// TIA Portal project "Sistema_de_silos" (V16) (continued)
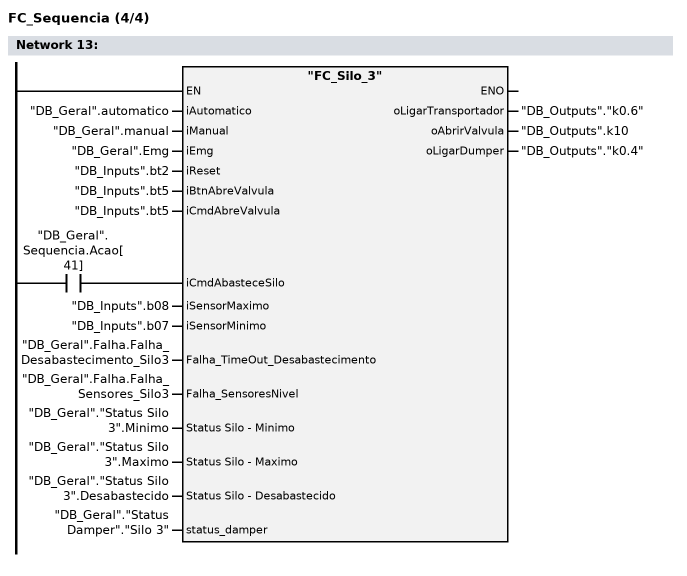
   RUNG wire#powerrail
      "FC_Silo_3"(iCmdAbasteceSilo := wire#w1, iAutomatico := "DB_Geral".automatico, iManual := "DB_Geral".manual, iEmg := "DB_Geral".Emg, iReset := "DB_Inputs".bt2, iBtnAbreValvula := "DB_Inputs".bt5, iCmdAbreValvula := "DB_Inputs".bt5, iSensorMaximo := "DB_Inputs".b08, iSensorMinimo := "DB_Inputs".b07, Falha_TimeOut_Desabastecimento := "DB_Geral".Falha.Falha_Desabastecimento_Silo3, Falha_SensoresNivel := "DB_Geral".Falha.Falha_Sensores_Silo3, "Status Silo - Minimo" := "DB_Geral"."Status Silo 3".Minimo, "Status Silo - Maximo" := "DB_Geral"."Status Silo 3".Maximo, "Status Silo - Desabastecido" := "DB_Geral"."Status Silo 3".Desabastecido, status_damper := "DB_Geral"."Status Damper"."Silo 3", oLigarTransportador => "DB_Outputs"."k0.6", oAbrirValvula => "DB_Outputs".k10, oLigarDumper => "DB_Outputs"."k0.4")
   END_RUNG
   RUNG wire#powerrail
      Contact( "DB_Geral".Sequencia.Acao[41] )
   END_RUNG wire#w1
   // the same network as SCL:
   "FC_Silo_3"(iAutomatico := "DB_Geral".automatico,
               iManual := "DB_Geral".manual,
               iEmg := "DB_Geral".Emg,
               iReset := "DB_Inputs".bt2,
               iBtnAbreValvula := "DB_Inputs".bt5,
               iCmdAbreValvula := "DB_Inputs".bt5,
               iCmdAbasteceSilo := "DB_Geral".Sequencia.Acao[41],
               iSensorMaximo := "DB_Inputs".b08,
               iSensorMinimo := "DB_Inputs".b07,
               Falha_TimeOut_Desabastecimento := "DB_Geral".Falha.Falha_Desabastecimento_Silo3,
               Falha_SensoresNivel := "DB_Geral".Falha.Falha_Sensores_Silo3,
               "Status Silo - Minimo" := "DB_Geral"."Status Silo 3".Minimo,
               "Status Silo - Maximo" := "DB_Geral"."Status Silo 3".Maximo,
               "Status Silo - Desabastecido" := "DB_Geral"."Status Silo 3".Desabastecido,
               status_damper := "DB_Geral"."Status Damper"."Silo 3",
               oLigarTransportador => "DB_Outputs"."k0.6",
               oAbrirValvula => "DB_Outputs".k10,
               oLigarDumper => "DB_Outputs"."k0.4");
END_REGION
END_FUNCTION

FUNCTION "FC_Silo_2" : Void   // FC5, LAD
{ S7_Optimized_Access := 'TRUE' }
VERSION : 0.1
   VAR_INPUT
      iAutomatico : Bool;
      iManual : Bool;
      iEmg : Bool;
      iReset : Bool;
      iBtnAbreValvula : Bool;
      iCmdAbreValvula : Bool;
      iCmdAbasteceSilo : Bool;
      iSensorMaximo : Bool;
      iSensorMinimo : Bool;
   END_VAR
   VAR_OUTPUT
      oLigarTransportador : Bool;
      oAbrirValvula : Bool;
      oLigarDumper : Bool;
   END_VAR
   VAR_IN_OUT
      Falha_TimeOut_Desabastecimento : Bool;
      Falha_SensoresNivel : Bool;
      "Status Silo - Minimo" : Bool;
      "Status Silo - Maximo" : Bool;
      "Status Silo - Desabastecido" : Bool;
      status_damper : Bool;
   END_VAR
   VAR CONSTANT
      Velocidade_fluxo : Int := 12;
   END_VAR
BEGIN

REGION Network 1
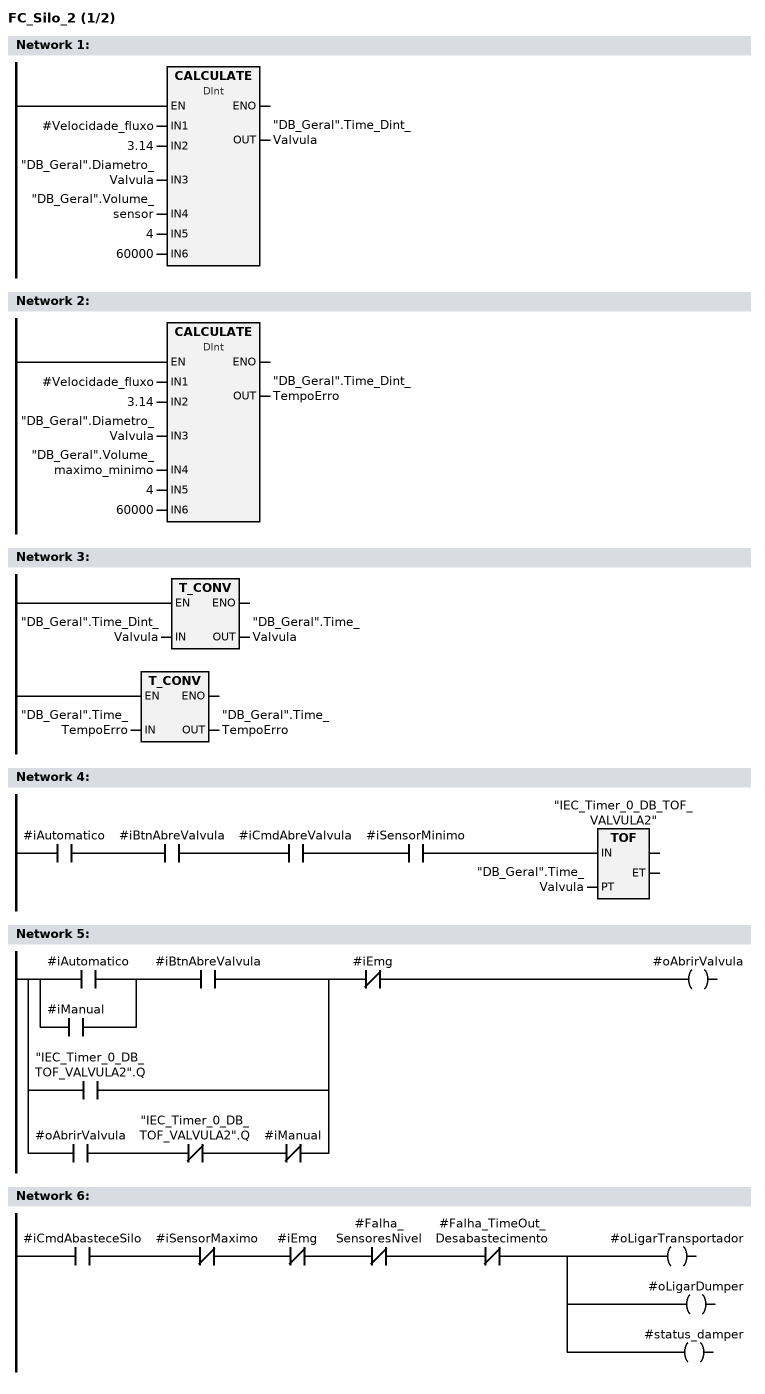
   RUNG wire#powerrail
      { S7_Templates := "SrcType := DInt"; S7_Expression := "(IN4 / (IN1* ((IN2*IN3*IN3) / IN5))) * IN6" } Calculate(in1 := #Velocidade_fluxo, in2 := 3.14, in3 := "DB_Geral".Diametro_Valvula, in4 := "DB_Geral".Volume_sensor, in5 := 4, in6 := 60000, out => "DB_Geral".Time_Dint_Valvula)
   END_RUNG
   // the same network as SCL:
   "DB_Geral".Time_Dint_Valvula := ("DB_Geral".Volume_sensor / (#Velocidade_fluxo* ((3.14*"DB_Geral".Diametro_Valvula*"DB_Geral".Diametro_Valvula) / 4))) * 60000;
END_REGION

REGION Network 2
   RUNG wire#powerrail
      { S7_Templates := "SrcType := DInt"; S7_Expression := "(IN4 / (IN1* ((IN2*IN3*IN3) / IN5))) * IN6" } Calculate(in1 := #Velocidade_fluxo, in2 := 3.14, in3 := "DB_Geral".Diametro_Valvula, in4 := "DB_Geral".Volume_maximo_minimo, in5 := 4, in6 := 60000, out => "DB_Geral".Time_Dint_TempoErro)
   END_RUNG
   // the same network as SCL:
   "DB_Geral".Time_Dint_TempoErro := ("DB_Geral".Volume_maximo_minimo / (#Velocidade_fluxo* ((3.14*"DB_Geral".Diametro_Valvula*"DB_Geral".Diametro_Valvula) / 4))) * 60000;
END_REGION

REGION Network 3
   "DB_Geral".Time_Valvula := T_CONV(IN := "DB_Geral".Time_Dint_Valvula);
   "DB_Geral".Time_TempoErro := T_CONV(IN := "DB_Geral".Time_TempoErro);
END_REGION

REGION Network 4
   "IEC_Timer_0_DB_TOF_VALVULA2".TOF(IN := #iAutomatico AND #iBtnAbreValvula AND #iCmdAbreValvula AND #iSensorMinimo,
                           PT := "DB_Geral".Time_Valvula);
END_REGION

REGION Network 5
   RUNG wire#powerrail
      Contact( #iAutomatico )
      wire#w1
      Contact( #iBtnAbreValvula )
      wire#w2
      I_Contact( #iEmg )
      Coil( #oAbrirValvula )
   END_RUNG
   RUNG wire#powerrail
      Contact( #iManual )
   END_RUNG wire#w1
   RUNG wire#powerrail
      Contact( "IEC_Timer_0_DB_TOF_VALVULA2".Q )
   END_RUNG wire#w2
   RUNG wire#powerrail
      Contact( #oAbrirValvula )
      I_Contact( "IEC_Timer_0_DB_TOF_VALVULA2".Q )
      I_Contact( #iManual )
   END_RUNG wire#w2
   // the same network as SCL:
   #oAbrirValvula := (((#iAutomatico OR #iManual) AND #iBtnAbreValvula) OR "IEC_Timer_0_DB_TOF_VALVULA2".Q OR (#oAbrirValvula AND NOT "IEC_Timer_0_DB_TOF_VALVULA2".Q AND NOT #iManual)) AND NOT #iEmg;
END_REGION

REGION Network 6
   RUNG wire#powerrail
      Contact( #iCmdAbasteceSilo )
      I_Contact( #iSensorMaximo )
      I_Contact( #iEmg )
      I_Contact( #Falha_SensoresNivel )
      I_Contact( #Falha_TimeOut_Desabastecimento )
      wire#w1
      Coil( #oLigarTransportador )
   END_RUNG
   RUNG wire#w1
      Coil( #oLigarDumper )
   END_RUNG
   RUNG wire#w1
      Coil( #status_damper )
   END_RUNG
   // the same network as SCL:
   #oLigarTransportador := #iCmdAbasteceSilo AND NOT #iSensorMaximo AND NOT #iEmg AND NOT #Falha_SensoresNivel AND NOT #Falha_TimeOut_Desabastecimento;
   #oLigarDumper := #oLigarTransportador;
   #status_damper := #oLigarTransportador;
END_REGION

REGION Network 7: Silo Principal - Reserva do produto
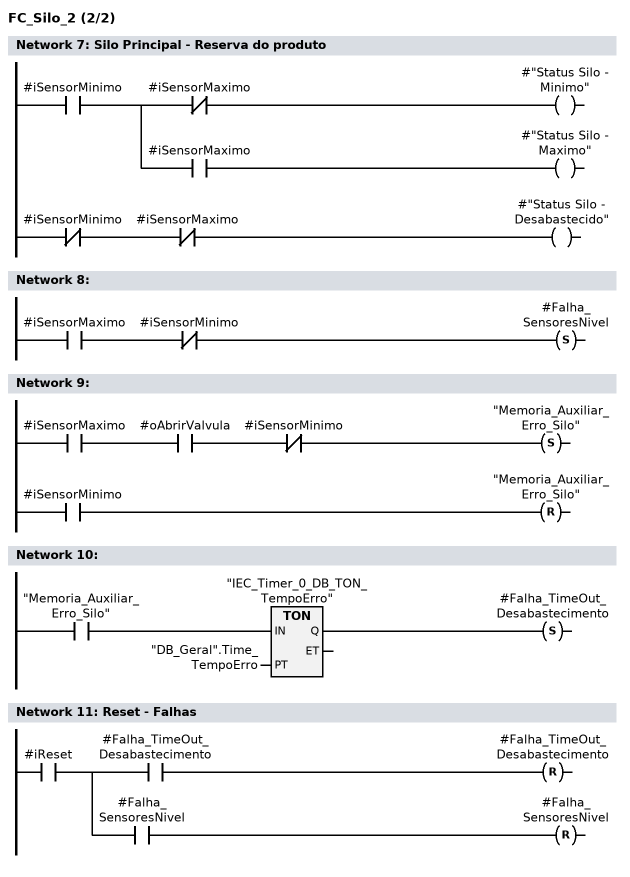
   RUNG wire#powerrail
      Contact( #iSensorMinimo )
      wire#w1
      I_Contact( #iSensorMaximo )
      Coil( #"Status Silo - Minimo" )
   END_RUNG
   RUNG wire#w1
      Contact( #iSensorMaximo )
      Coil( #"Status Silo - Maximo" )
   END_RUNG
   RUNG wire#powerrail
      I_Contact( #iSensorMinimo )
      I_Contact( #iSensorMaximo )
      Coil( #"Status Silo - Desabastecido" )
   END_RUNG
   // the same network as SCL:
   #"Status Silo - Minimo" := #iSensorMinimo AND NOT #iSensorMaximo;
   #"Status Silo - Maximo" := #iSensorMinimo AND #iSensorMaximo;
   #"Status Silo - Desabastecido" := NOT #iSensorMinimo AND NOT #iSensorMaximo;
END_REGION

REGION Network 8
   RUNG wire#powerrail
      Contact( #iSensorMaximo )
      I_Contact( #iSensorMinimo )
      S_Coil( #Falha_SensoresNivel )
   END_RUNG
   // the same network as SCL:
   IF #iSensorMaximo AND NOT #iSensorMinimo THEN #Falha_SensoresNivel := TRUE; END_IF;
END_REGION

REGION Network 9
   RUNG wire#powerrail
      Contact( #iSensorMaximo )
      Contact( #oAbrirValvula )
      I_Contact( #iSensorMinimo )
      S_Coil( "Memoria_Auxiliar_Erro_Silo" )
   END_RUNG
   RUNG wire#powerrail
      Contact( #iSensorMinimo )
      R_Coil( "Memoria_Auxiliar_Erro_Silo" )
   END_RUNG
   // the same network as SCL:
   IF #iSensorMaximo AND #oAbrirValvula AND NOT #iSensorMinimo THEN
       "Memoria_Auxiliar_Erro_Silo" := TRUE;
   END_IF;
   IF #iSensorMinimo THEN "Memoria_Auxiliar_Erro_Silo" := FALSE; END_IF;
END_REGION

REGION Network 10
   "IEC_Timer_0_DB_TON_TempoErro".TON(IN := "Memoria_Auxiliar_Erro_Silo", PT := "DB_Geral".Time_TempoErro);
   IF "IEC_Timer_0_DB_TON_TempoErro".Q THEN #Falha_TimeOut_Desabastecimento := TRUE; END_IF;
END_REGION

REGION Network 11: Reset - Falhas
   RUNG wire#powerrail
      Contact( #iReset )
      wire#w1
      Contact( #Falha_TimeOut_Desabastecimento )
      R_Coil( #Falha_TimeOut_Desabastecimento )
   END_RUNG
   RUNG wire#w1
      Contact( #Falha_SensoresNivel )
      R_Coil( #Falha_SensoresNivel )
   END_RUNG
   // the same network as SCL:
   IF #iReset AND #Falha_TimeOut_Desabastecimento THEN #Falha_TimeOut_Desabastecimento := FALSE; END_IF;
   IF #iReset AND #Falha_SensoresNivel THEN #Falha_SensoresNivel := FALSE; END_IF;
END_REGION
END_FUNCTION

FUNCTION "FC_Silo_Principal" : Void   // FC6, LAD
{ S7_Optimized_Access := 'TRUE' }
VERSION : 0.1
   VAR_INPUT
      iAutomatico : Bool;
      iManual : Bool;
      iEmg : Bool;
      iReset : Bool;
      iBtnAbasteceSilo : Bool;
      iCmdAbasteceSilo : Bool;
      iSensorMaximo : Bool;
      iSensorMinimo : Bool;
   END_VAR
   VAR_OUTPUT
      oAbasteceSilo : Bool;
   END_VAR
   VAR_IN_OUT
      Falha_SensoresNivel : Bool;
      "Status Silo - Minimo" : Bool;
      "Status Silo - Maximo" : Bool;
      "Status Silo - Desabastecido" : Bool;
   END_VAR
BEGIN

REGION Network 1
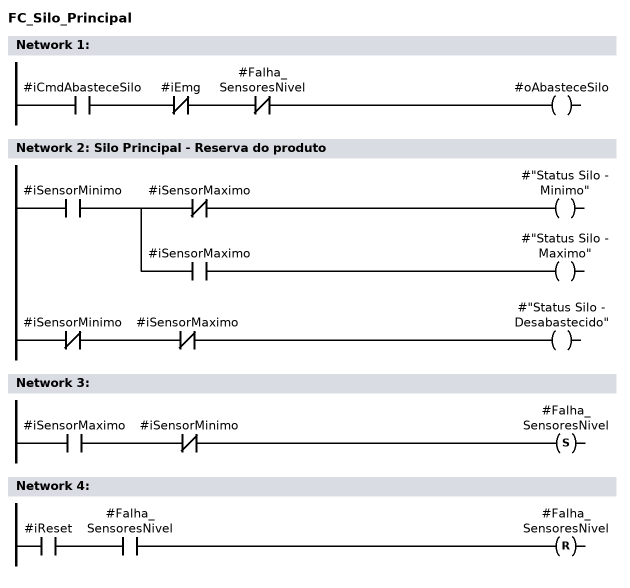
   RUNG wire#powerrail
      Contact( #iCmdAbasteceSilo )
      I_Contact( #iEmg )
      I_Contact( #Falha_SensoresNivel )
      Coil( #oAbasteceSilo )
   END_RUNG
   // the same network as SCL:
   #oAbasteceSilo := #iCmdAbasteceSilo AND NOT #iEmg AND NOT #Falha_SensoresNivel;
END_REGION

REGION Network 2: Silo Principal - Reserva do produto
   RUNG wire#powerrail
      Contact( #iSensorMinimo )
      wire#w1
      I_Contact( #iSensorMaximo )
      Coil( #"Status Silo - Minimo" )
   END_RUNG
   RUNG wire#w1
      Contact( #iSensorMaximo )
      Coil( #"Status Silo - Maximo" )
   END_RUNG
   RUNG wire#powerrail
      I_Contact( #iSensorMinimo )
      I_Contact( #iSensorMaximo )
      Coil( #"Status Silo - Desabastecido" )
   END_RUNG
   // the same network as SCL:
   #"Status Silo - Minimo" := #iSensorMinimo AND NOT #iSensorMaximo;
   #"Status Silo - Maximo" := #iSensorMinimo AND #iSensorMaximo;
   #"Status Silo - Desabastecido" := NOT #iSensorMinimo AND NOT #iSensorMaximo;
END_REGION

REGION Network 3
   RUNG wire#powerrail
      Contact( #iSensorMaximo )
      I_Contact( #iSensorMinimo )
      S_Coil( #Falha_SensoresNivel )
   END_RUNG
   // the same network as SCL:
   IF #iSensorMaximo AND NOT #iSensorMinimo THEN #Falha_SensoresNivel := TRUE; END_IF;
END_REGION

REGION Network 4
   RUNG wire#powerrail
      Contact( #iReset )
      Contact( #Falha_SensoresNivel )
      R_Coil( #Falha_SensoresNivel )
   END_RUNG
   // the same network as SCL:
   IF #iReset AND #Falha_SensoresNivel THEN #Falha_SensoresNivel := FALSE; END_IF;
END_REGION
END_FUNCTION

FUNCTION "FC_Silo_3" : Void   // FC7, LAD
{ S7_Optimized_Access := 'TRUE' }
VERSION : 0.1
   VAR_INPUT
      iAutomatico : Bool;
      iManual : Bool;
      iEmg : Bool;
      iReset : Bool;
      iBtnAbreValvula : Bool;
      iCmdAbreValvula : Bool;
      iCmdAbasteceSilo : Bool;
      iSensorMaximo : Bool;
      iSensorMinimo : Bool;
   END_VAR
   VAR_OUTPUT
      oLigarTransportador : Bool;
      oAbrirValvula : Bool;
      oLigarDumper : Bool;
   END_VAR
   VAR_IN_OUT
      Falha_TimeOut_Desabastecimento : Bool;
      Falha_SensoresNivel : Bool;
      "Status Silo - Minimo" : Bool;
      "Status Silo - Maximo" : Bool;
      "Status Silo - Desabastecido" : Bool;
      status_damper : Bool;
   END_VAR
   VAR CONSTANT
      Velocidade_fluxo : Int := 12;
   END_VAR
BEGIN

REGION Network 1
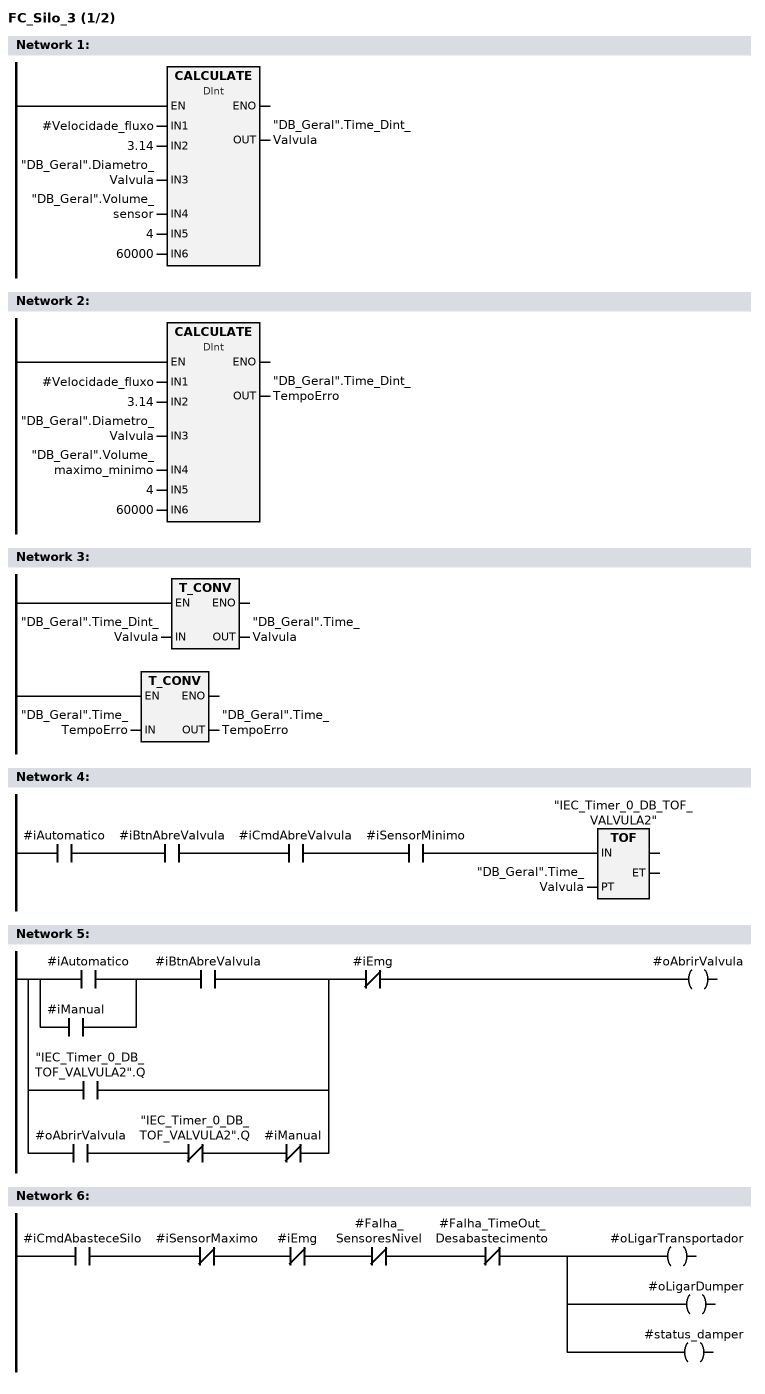
   RUNG wire#powerrail
      { S7_Templates := "SrcType := DInt"; S7_Expression := "(IN4 / (IN1* ((IN2*IN3*IN3) / IN5))) * IN6" } Calculate(in1 := #Velocidade_fluxo, in2 := 3.14, in3 := "DB_Geral".Diametro_Valvula, in4 := "DB_Geral".Volume_sensor, in5 := 4, in6 := 60000, out => "DB_Geral".Time_Dint_Valvula)
   END_RUNG
   // the same network as SCL:
   "DB_Geral".Time_Dint_Valvula := ("DB_Geral".Volume_sensor / (#Velocidade_fluxo* ((3.14*"DB_Geral".Diametro_Valvula*"DB_Geral".Diametro_Valvula) / 4))) * 60000;
END_REGION

REGION Network 2
   RUNG wire#powerrail
      { S7_Templates := "SrcType := DInt"; S7_Expression := "(IN4 / (IN1* ((IN2*IN3*IN3) / IN5))) * IN6" } Calculate(in1 := #Velocidade_fluxo, in2 := 3.14, in3 := "DB_Geral".Diametro_Valvula, in4 := "DB_Geral".Volume_maximo_minimo, in5 := 4, in6 := 60000, out => "DB_Geral".Time_Dint_TempoErro)
   END_RUNG
   // the same network as SCL:
   "DB_Geral".Time_Dint_TempoErro := ("DB_Geral".Volume_maximo_minimo / (#Velocidade_fluxo* ((3.14*"DB_Geral".Diametro_Valvula*"DB_Geral".Diametro_Valvula) / 4))) * 60000;
END_REGION

REGION Network 3
   "DB_Geral".Time_Valvula := T_CONV(IN := "DB_Geral".Time_Dint_Valvula);
   "DB_Geral".Time_TempoErro := T_CONV(IN := "DB_Geral".Time_TempoErro);
END_REGION

REGION Network 4
   "IEC_Timer_0_DB_TOF_VALVULA2".TOF(IN := #iAutomatico AND #iBtnAbreValvula AND #iCmdAbreValvula AND #iSensorMinimo,
                           PT := "DB_Geral".Time_Valvula);
END_REGION

REGION Network 5
   RUNG wire#powerrail
      Contact( #iAutomatico )
      wire#w1
      Contact( #iBtnAbreValvula )
      wire#w2
      I_Contact( #iEmg )
      Coil( #oAbrirValvula )
   END_RUNG
   RUNG wire#powerrail
      Contact( #iManual )
   END_RUNG wire#w1
   RUNG wire#powerrail
      Contact( "IEC_Timer_0_DB_TOF_VALVULA2".Q )
   END_RUNG wire#w2
   RUNG wire#powerrail
      Contact( #oAbrirValvula )
      I_Contact( "IEC_Timer_0_DB_TOF_VALVULA2".Q )
      I_Contact( #iManual )
   END_RUNG wire#w2
   // the same network as SCL:
   #oAbrirValvula := (((#iAutomatico OR #iManual) AND #iBtnAbreValvula) OR "IEC_Timer_0_DB_TOF_VALVULA2".Q OR (#oAbrirValvula AND NOT "IEC_Timer_0_DB_TOF_VALVULA2".Q AND NOT #iManual)) AND NOT #iEmg;
END_REGION

REGION Network 6
   RUNG wire#powerrail
      Contact( #iCmdAbasteceSilo )
      I_Contact( #iSensorMaximo )
      I_Contact( #iEmg )
      I_Contact( #Falha_SensoresNivel )
      I_Contact( #Falha_TimeOut_Desabastecimento )
      wire#w1
      Coil( #oLigarTransportador )
   END_RUNG
   RUNG wire#w1
      Coil( #oLigarDumper )
   END_RUNG
   RUNG wire#w1
      Coil( #status_damper )
   END_RUNG
   // the same network as SCL:
   #oLigarTransportador := #iCmdAbasteceSilo AND NOT #iSensorMaximo AND NOT #iEmg AND NOT #Falha_SensoresNivel AND NOT #Falha_TimeOut_Desabastecimento;
   #oLigarDumper := #oLigarTransportador;
   #status_damper := #oLigarTransportador;
END_REGION

REGION Network 7: Silo Principal - Reserva do produto
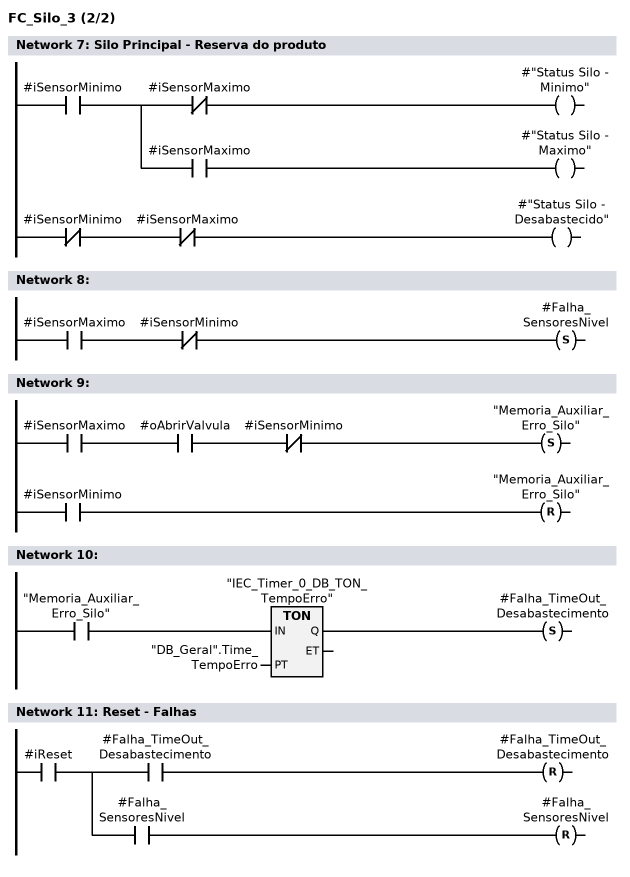
   RUNG wire#powerrail
      Contact( #iSensorMinimo )
      wire#w1
      I_Contact( #iSensorMaximo )
      Coil( #"Status Silo - Minimo" )
   END_RUNG
   RUNG wire#w1
      Contact( #iSensorMaximo )
      Coil( #"Status Silo - Maximo" )
   END_RUNG
   RUNG wire#powerrail
      I_Contact( #iSensorMinimo )
      I_Contact( #iSensorMaximo )
      Coil( #"Status Silo - Desabastecido" )
   END_RUNG
   // the same network as SCL:
   #"Status Silo - Minimo" := #iSensorMinimo AND NOT #iSensorMaximo;
   #"Status Silo - Maximo" := #iSensorMinimo AND #iSensorMaximo;
   #"Status Silo - Desabastecido" := NOT #iSensorMinimo AND NOT #iSensorMaximo;
END_REGION

REGION Network 8
   RUNG wire#powerrail
      Contact( #iSensorMaximo )
      I_Contact( #iSensorMinimo )
      S_Coil( #Falha_SensoresNivel )
   END_RUNG
   // the same network as SCL:
   IF #iSensorMaximo AND NOT #iSensorMinimo THEN #Falha_SensoresNivel := TRUE; END_IF;
END_REGION

REGION Network 9
   RUNG wire#powerrail
      Contact( #iSensorMaximo )
      Contact( #oAbrirValvula )
      I_Contact( #iSensorMinimo )
      S_Coil( "Memoria_Auxiliar_Erro_Silo" )
   END_RUNG
   RUNG wire#powerrail
      Contact( #iSensorMinimo )
      R_Coil( "Memoria_Auxiliar_Erro_Silo" )
   END_RUNG
   // the same network as SCL:
   IF #iSensorMaximo AND #oAbrirValvula AND NOT #iSensorMinimo THEN
       "Memoria_Auxiliar_Erro_Silo" := TRUE;
   END_IF;
   IF #iSensorMinimo THEN "Memoria_Auxiliar_Erro_Silo" := FALSE; END_IF;
END_REGION

REGION Network 10
   "IEC_Timer_0_DB_TON_TempoErro".TON(IN := "Memoria_Auxiliar_Erro_Silo", PT := "DB_Geral".Time_TempoErro);
   IF "IEC_Timer_0_DB_TON_TempoErro".Q THEN #Falha_TimeOut_Desabastecimento := TRUE; END_IF;
END_REGION

REGION Network 11: Reset - Falhas
   RUNG wire#powerrail
      Contact( #iReset )
      wire#w1
      Contact( #Falha_TimeOut_Desabastecimento )
      R_Coil( #Falha_TimeOut_Desabastecimento )
   END_RUNG
   RUNG wire#w1
      Contact( #Falha_SensoresNivel )
      R_Coil( #Falha_SensoresNivel )
   END_RUNG
   // the same network as SCL:
   IF #iReset AND #Falha_TimeOut_Desabastecimento THEN #Falha_TimeOut_Desabastecimento := FALSE; END_IF;
   IF #iReset AND #Falha_SensoresNivel THEN #Falha_SensoresNivel := FALSE; END_IF;
END_REGION
END_FUNCTION

ORGANIZATION_BLOCK "Main"   // OB1, LAD, ProgramCycle
TITLE = "Main Program Sweep (Cycle)"
{ S7_Optimized_Access := 'TRUE' }
VERSION : 0.1
   VAR_INPUT
      Initial_Call : Bool;   // Initial call of this OB
      Remanence : Bool;   // =True, if remanent data are available
   END_VAR
BEGIN

REGION Network 1
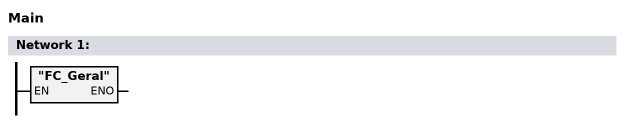
   RUNG wire#powerrail
      "FC_Geral"()
   END_RUNG
   // the same network as SCL:
   "FC_Geral"();
END_REGION
END_ORGANIZATION_BLOCK

(* ===== HMI "HMI_RT_1" =====
system functions are stored by id; their names below are inferred from use
connection "HMI_Connection_2": ETHERNET, S7_1200_OMS

HMI tags "Default tag table"
   "Tag_ScreenNumber" : UInt, internal
   "bt1" : Bool = PLC bt1 AT %I0.1, 1 s
   "bt0" : Bool = PLC bt0 AT %I0.0, 1 s
   "bt3" : Bool = PLC bt3 AT %I0.3, 1 s
   "bt2" : Bool = PLC bt2 AT %I0.2, 1 s
   "DB_Inputs_bt1" : Bool = PLC DB_Inputs.bt1, 1 s
   "DB_Inputs_bt0" : Bool = PLC DB_Inputs.bt0, 1 s
   "DB_Inputs_bt3" : Bool = PLC DB_Inputs.bt3, 1 s
   "DB_Inputs_bt2" : Bool = PLC DB_Inputs.bt2, 1 s
   "DB_Inputs_bt4" : Bool = PLC DB_Inputs.bt4, 1 s
   "DB_Inputs_bt5" : Bool = PLC DB_Inputs.bt5, 1 s
   "DB_Inputs_b04" : Bool = PLC DB_Inputs.b04, 1 s
   "DB_Inputs_b03" : Bool = PLC DB_Inputs.b03, 1 s
   "DB_Outputs_k0.5" : Bool = PLC DB_Outputs."k0.5", 1 s
   "DB_Outputs_k0.6" : Bool = PLC DB_Outputs."k0.6", 1 s
   "DB_Outputs_k0.7" : Bool = PLC DB_Outputs."k0.7", 1 s
   "DB_Geral_Falha_Falha_Desabastecimento_Silo2" : Bool = PLC DB_Geral.Falha.Falha_Desabastecimento_Silo2, 1 s
   "DB_Outputs_k10" : Bool = PLC DB_Outputs.k10, 1 s
   "DB_Geral_Falha_Falha_Desabastecimento_Silo3" : Bool = PLC DB_Geral.Falha.Falha_Desabastecimento_Silo3, 1 s
   "DB_Inputs_b01" : Bool = PLC DB_Inputs.b01, 1 s
   "DB_Geral_Falha_Falha_Sensores_SiloPrincipal" : Bool = PLC DB_Geral.Falha.Falha_Sensores_SiloPrincipal, 1 s
   "DB_Inputs_b02" : Bool = PLC DB_Inputs.b02, 1 s
   "DB_Geral_Falha_Falha_Sensores_Silo2" : Bool = PLC DB_Geral.Falha.Falha_Sensores_Silo2, 1 s
   "DB_Inputs_b05" : Bool = PLC DB_Inputs.b05, 1 s
   "DB_Inputs_b06" : Bool = PLC DB_Inputs.b06, 1 s
   "DB_Geral_Falha_Falha_Sensores_Silo3" : Bool = PLC DB_Geral.Falha.Falha_Sensores_Silo3, 1 s
   "DB_Inputs_b07" : Bool = PLC DB_Inputs.b07, 1 s
   "DB_Inputs_b08" : Bool = PLC DB_Inputs.b08, 1 s
   "DB_Geral_Status Damper_Ligado" : Bool = PLC DB_Geral."Status Damper".Ligado, 1 s
   "DB_Geral_Status Damper_Silo 2" : Bool = PLC DB_Geral."Status Damper"."Silo 2", 1 s
   "DB_Geral_Status Damper_Silo 3" : Bool = PLC DB_Geral."Status Damper"."Silo 3", 1 s
   "DB_Geral_number_status" : Int = PLC DB_Geral.number_status, 1 s
   "DB_Geral_automatico" : Bool = PLC DB_Geral.automatico, 1 s
   "DB_Geral_manual" : Bool = PLC DB_Geral.manual, 1 s

HMI tags "Animation"
   "Tag_op" : Bool, internal

graphic list "sensor_damper_silo3Aberto": 0 'Group 1000005174'; 1 'sensor_silo3_damper_aberto'

graphic list "sensor_damper_silo2Aberto": 0 'Group 1000005187'; 1 'sensor_silo2_damper_aberto_acionado'

graphic list "transportador": 0 'conveyor'; 1 'transportador_acionado'

graphic list "sensores_nivel": 0 'Sensores_nivel_normal_1'; 1 'sensores_nivel_acionado'

graphic list "valvula2": 0 'valvula2'; 1 'valvula2_acionada'

graphic list "valvula3": 0 'Valvula3'; 1 'Valvula3_acionada'

graphic list "damper2": 0 'damper_desligado'; 1 'damper_silo2_acionado'

graphic list "damper3": 0 'damper_desligado'; 1 'damper_silo3_acionado'

graphic list "sensores_nivel_falha": 0 ''; 1 'Sensores_nivel_falha_1'

graphic list "valvula2_Falha": 0 ''; 1 'valvula2_falha'

graphic list "valvula3_falha": 0 ''; 1 'Valvula3_falha'

graphic list "Status": 0 'StatusManual'; 1 'statusAutomatico'; 2 'StatusEmg'; 3 'statusFalha'; 4 'statusSemModo'

graphic list "manual": 0 'StatusManual_off'; 1 'StatusManual'

graphic list "automatico": 0 'statusAutomatico_off'; 1 'statusAutomatico'

graphic list "emergencia": 1 'StatusEmg_off'; 0 'StatusEmg'

graphic list "reset": 0 'statusSemModo_off'; 1 'Reset'

graphic list "btn_valvula2": 0 'btn_valv2off_1'; 1 'btn_val3'

graphic list "btn_valvula3": 0 'btn_val3off'; 1 'btn_val2_1'

screen "Root screen" 1280x740, template "Template_1"
   on GenerateScreen: SetTag("Tag_ScreenNumber", 1)
   Button "HmiScreenItemData" at 79,35 size 213x73; TextOff 'Teste Screen'; PictureOff "Navigates to Teste Screen for TP1200 Comfort 16.0.0.0"; PictureOn "Navigates to Teste Screen for TP1200 Comfort 16.0.0.0"
      on Release: ActivateScreen("Teste Screen", 0)
   Button "HmiScreenItemData_1" at 1002,36 size 213x73; TextOff 'Operation Screen'; PictureOff "Navigates to Operation Screen for TP1200 Comfort 16.0.0.0"; PictureOn "Navigates to Operation Screen for TP1200 Comfort 16.0.0.0"
      on Release: ActivateScreen("Operation Screen", 0)
   Button "HmiScreenItemData_2" at 692,33 size 213x73; TextOff 'Fail/Emg Screen'; PictureOff "Navigates to Fail/Emg Screen for TP1200 Comfort 16.0.0.0"; PictureOn "Navigates to Fail/Emg Screen for TP1200 Comfort 16.0.0.0"
      on Release: ActivateScreen("Fail/Emg Screen", 0)
   Button "HmiScreenItemData_4" at 377,35 size 213x73; TextOff 'System screens'; PictureOff "Navigates to System screens for TP1200 Comfort 16.0.0.0"; PictureOn "Navigates to System screens for TP1200 Comfort 16.0.0.0"
      on Release: ActivateScreen("System screens", 0)
   GraphicView "Graphic view_3" at 361,257 size 541x174; Picture "Siemens Logo"

Template "Template_1" 1280x740
   Button "Exit" at 1200,679 size 78x59; TextOff 'Exit'; PictureOff "ExitRuntime_TP1200_Comfort_TR"; PictureOn "ExitRuntime_TP1200_Comfort_TR"
      on Release: StopRuntime(0)
   Button "Template_Button" at 1120,679 size 78x59; TextOff 'Text'
   Button "Template_Button_1" at 1040,679 size 78x59; TextOff 'Text'
   Button "Template_Button_2" at 960,679 size 78x59; TextOff 'Text'
   Button "Template_Button_3" at 880,679 size 78x59; TextOff 'Text'
   Button "Template_Button_4" at 800,679 size 78x59; TextOff 'Text'
   Button "Template_Button_5" at 720,679 size 78x59; TextOff 'Text'
   Button "Template_Button_6" at 640,679 size 78x59; TextOff 'Text'
   Button "Template_Button_7" at 561,679 size 78x59; TextOff 'Text'
   Button "Template_Button_8" at 481,679 size 78x59; TextOff 'Text'
   Button "Template_Button_9" at 401,679 size 78x59; TextOff 'Text'
   Button "Template_Button_10" at 321,679 size 78x59; TextOff 'Text'
   Button "Template_Button_11" at 241,679 size 78x59; TextOff 'Text'
   Button "Template_Button_12" at 161,679 size 78x59; TextOff 'Text'
   Button "Alarms" at 81,679 size 78x59; TextOff 'Alarms'; PictureOff "AlarmDisplay_TP1200_Comfort_TR"; PictureOn "AlarmDisplay_TP1200_Comfort_TR"
      on Release: function_ef3f5d25("Alarm window_Unacknowledged", -1)
   Button "Start screen" at 1,679 size 78x59; TextOff 'Start screen'; PictureOff "NavigateHome_TP1200_Comfort_TR"; PictureOn "NavigateHome_TP1200_Comfort_TR"
      on Release: ActivateScreen("Root screen", 0)

screen "Teste Screen" 1280x740, template "Template_1"
   on GenerateScreen: SetTag("Tag_ScreenNumber", 2)
   Rectangle "Rectangle_1" at 0,130 size 201x292
      Visibility <- "Tag_op"
   Button "Button_1" at 14,140 size 173x52; TextOff 'Text'; PictureOff "StatusManual"; PictureList "manual"
      Visibility <- "Tag_op"
      on Press: InvertBit("DB_Inputs_bt1")
      ProcessValue <- "DB_Inputs_bt1"
   Button "Button_2" at 14,213 size 173x52; TextOff 'Text'; PictureOff "statusAutomatico"; PictureList "automatico"
      Visibility <- "Tag_op"
      on Press: InvertBit("DB_Inputs_bt0")
      ProcessValue <- "DB_Inputs_bt0"
   Button "Button_3" at 14,285 size 173x52; TextOff 'Text'; PictureOff "StatusEmg"; PictureList "emergencia"
      Visibility <- "Tag_op"
      on Press: InvertBit("DB_Inputs_bt3")
      ProcessValue <- "DB_Inputs_bt3"
   Button "Button_4" at 14,357 size 173x52; TextOff 'Text'; PictureOff "Reset"; PictureList "reset"
      Visibility <- "Tag_op"
      on Press: InvertBit("DB_Inputs_bt2")
      ProcessValue <- "DB_Inputs_bt2"
   Rectangle "Rectangle_2" at 0,436 size 202x143
      Visibility <- "Tag_op"
   Button "Back" at 0,0 size 112x36; TextOff 'Back'
      on Release: ActivateScreen("Root screen", 0)
   GraphicView "Graphic view_6" at 697,48 size 165x302; Picture "Clip_path_group_1-removebg-preview"
   Button "Button_5" at 14,515 size 179x56; TextOff 'Text'; PictureOff "btn_val2_1"; PictureList "btn_valvula3"
      Visibility <- "Tag_op"
      on Click: InvertBit("DB_Inputs_bt4")
      ProcessValue <- "DB_Inputs_bt5"
   Button "Button_6" at 13,445 size 179x56; TextOff 'Text'; PictureOff "btn_val3"; PictureList "btn_valvula2"
      Visibility <- "Tag_op"
      on Click: InvertBit("DB_Inputs_bt5")
      ProcessValue <- "DB_Inputs_bt4"
   Group "Group_2" at 0,130 size 201x292; PictureOff "StatusManual"
   Button "Button_7" at 0,93 size 199x32; TextOff 'Operação'
      on Click: InvertBit("Tag_op")
   GraphicIOField "Graphic I/O field_1" at 717,246 size 41x16; PictureList "sensor_damper_silo3Aberto"
      ProcessValue <- "DB_Inputs_b04"
   GraphicIOField "Graphic I/O field_2" at 808,245 size 41x16; PictureList "sensor_damper_silo2Aberto"
      ProcessValue <- "DB_Inputs_b03"
   GraphicIOField "Graphic I/O field_3" at 567,372 size 178x32; PictureList "transportador"
      ProcessValue <- "DB_Outputs_k0.5"
   GraphicIOField "Graphic I/O field_4" at 823,371 size 178x32; PictureList "transportador"
      ProcessValue <- "DB_Outputs_k0.6"
   GraphicView "Graphic view_3" at 438,415 size 126x229; Picture "silo2"
   GraphicIOField "Graphic I/O field_5" at 388,623 size 96x20; PictureList "valvula2"
      ProcessValue <- "DB_Outputs_k0.7"
      Visibility <- "DB_Geral_Falha_Falha_Desabastecimento_Silo2"
   GraphicView "Graphic view_5" at 992,415 size 126x228; Picture "silo2"
   GraphicIOField "Graphic I/O field_6" at 1073,623 size 96x20; PictureList "valvula3"
      ProcessValue <- "DB_Outputs_k10"
      Visibility <- "DB_Geral_Falha_Falha_Desabastecimento_Silo3"
   GraphicIOField "Graphic I/O field_7" at 388,623 size 96x20; PictureList "valvula2_Falha"
      Visibility <- "DB_Geral_Falha_Falha_Desabastecimento_Silo2"
      ProcessValue <- "DB_Geral_Falha_Falha_Desabastecimento_Silo2"
   GraphicIOField "Graphic I/O field_8" at 1073,623 size 96x20; PictureList "valvula3_falha"
      Visibility <- "DB_Geral_Falha_Falha_Desabastecimento_Silo3"
      ProcessValue <- "DB_Geral_Falha_Falha_Desabastecimento_Silo3"
   GraphicIOField "Graphic I/O field_9" at 638,58 size 305x23; PictureList "sensores_nivel"
      Visibility <- "DB_Geral_Falha_Falha_Sensores_SiloPrincipal"
      ProcessValue <- "DB_Inputs_b02"
   GraphicIOField "Graphic I/O field_10" at 641,166 size 305x23; PictureList "sensores_nivel"
      Visibility <- "DB_Geral_Falha_Falha_Sensores_SiloPrincipal"
      ProcessValue <- "DB_Inputs_b01"
   GraphicIOField "Graphic I/O field_11" at 638,58 size 305x23; PictureList "sensores_nivel_falha"
      Visibility <- "DB_Geral_Falha_Falha_Sensores_SiloPrincipal"
      ProcessValue <- "DB_Geral_Falha_Falha_Sensores_SiloPrincipal"
   GraphicIOField "Graphic I/O field_12" at 641,166 size 305x23; PictureList "sensores_nivel_falha"
      ProcessValue <- "DB_Geral_Falha_Falha_Sensores_SiloPrincipal"
      Visibility <- "DB_Geral_Falha_Falha_Sensores_SiloPrincipal"
   GraphicIOField "Graphic I/O field_13" at 378,519 size 238x23; PictureList "sensores_nivel"
      ProcessValue <- "DB_Inputs_b05"
      Visibility <- "DB_Geral_Falha_Falha_Sensores_Silo2"
   GraphicIOField "Graphic I/O field_14" at 378,519 size 238x23; PictureList "sensores_nivel_falha"
      ProcessValue <- "DB_Geral_Falha_Falha_Sensores_Silo2"
      Visibility <- "DB_Geral_Falha_Falha_Sensores_Silo2"
   GraphicIOField "Graphic I/O field_15" at 378,420 size 238x23; PictureList "sensores_nivel"
      ProcessValue <- "DB_Inputs_b06"
      Visibility <- "DB_Geral_Falha_Falha_Sensores_Silo2"
   GraphicIOField "Graphic I/O field_16" at 378,420 size 238x23; PictureList "sensores_nivel_falha"
      Visibility <- "DB_Geral_Falha_Falha_Sensores_Silo2"
      ProcessValue <- "DB_Geral_Falha_Falha_Sensores_Silo2"
   GraphicIOField "Graphic I/O field_17" at 937,519 size 238x23; PictureList "sensores_nivel"
      ProcessValue <- "DB_Inputs_b07"
      Visibility <- "DB_Geral_Falha_Falha_Desabastecimento_Silo3"
   GraphicIOField "Graphic I/O field_18" at 937,519 size 238x23; PictureList "sensores_nivel_falha"
      Visibility <- "DB_Geral_Falha_Falha_Sensores_Silo3"
      ProcessValue <- "DB_Geral_Falha_Falha_Sensores_Silo3"
   GraphicIOField "Graphic I/O field_19" at 935,420 size 238x23; PictureList "sensores_nivel"
      Visibility <- "DB_Geral_Falha_Falha_Sensores_Silo3"
      ProcessValue <- "DB_Inputs_b08"
   GraphicIOField "Graphic I/O field_20" at 935,420 size 238x23; PictureList "sensores_nivel_falha"
      ProcessValue <- "DB_Geral_Falha_Falha_Sensores_Silo3"
      Visibility <- "DB_Geral_Falha_Falha_Sensores_Silo3"
   Button "Button_9" at 367,412 size 55x34; TextOff 'Text'
      on Press: InvertBit("DB_Inputs_b06")
   Button "Button_10" at 369,519 size 55x34; TextOff 'Text'
      on Press: InvertBit("DB_Inputs_b05")
   Button "Button_11" at 928,414 size 55x34; TextOff 'Text'
      on Press: InvertBit("DB_Inputs_b08")
   Button "Button_12" at 928,514 size 55x34; TextOff 'Text'
      on Press: InvertBit("DB_Inputs_b07")
   Button "Button_13" at 637,162 size 55x34; TextOff 'Text'
      on Press: InvertBit("DB_Inputs_b01")
   Button "Button_16" at 633,55 size 55x34; TextOff 'Text'
      on Press: InvertBit("DB_Inputs_b02")
   GraphicIOField "Graphic I/O field_21" at 754,245 size 60x22; PictureList "damper2"
      ProcessValue <- "DB_Geral_Status Damper_Silo 2"
      Visibility <- "DB_Geral_Status Damper_Silo 3"
   GraphicIOField "Graphic I/O field_22" at 754,244 size 60x22; PictureList "damper3"
      ProcessValue <- "DB_Geral_Status Damper_Silo 3"
      Visibility <- "DB_Geral_Status Damper_Silo 2"

screen "Operation Screen" 1280x740, template "Template_1"
   on GenerateScreen: SetTag("Tag_ScreenNumber", 3)
   TextField "HmiScreenItemData" at 128,324 size 1024x27; Text 'Operation Screen'
   Button "Back" at 1,1 size 159x47; TextOff 'Back'
      on Release: ActivateScreen("Root screen", 0)

screen "Fail/Emg Screen" 1280x740, template "Template_1"
   on GenerateScreen: SetTag("Tag_ScreenNumber", 4)
   TextField "HmiScreenItemData" at 128,324 size 1024x27; Text 'Fail/Emg Screen'
   Button "Back" at 1,1 size 159x47; TextOff 'Back'
      on Release: ActivateScreen("Root screen", 0)

screen "System screens" 1280x740, template "Template_1"
   on GenerateScreen: SetTag("Tag_ScreenNumber", 5)
   Button "Back" at 1,1 size 159x47; TextOff 'Back'
      on Release: ActivateScreen("Root screen", 0)
   Button "HmiScreenItemData" at 36,95 size 159x47; TextOff 'SIMATIC PLC system diagnos...'; PictureOff "Navigates to SIMATIC PLC system diagnostics for TP1200 Comfort 16.0.0.0"; PictureOn "Navigates to SIMATIC PLC system diagnostics for TP1200 Comfort 16.0.0.0"
      on Release: ActivateScreen("SIMATIC PLC system diagnostics", 0)
   Button "HmiScreenItemData_1" at 36,154 size 159x47; TextOff 'System settings'; PictureOff "Navigates to System settings for TP1200 Comfort 16.0.0.0"; PictureOn "Navigates to System settings for TP1200 Comfort 16.0.0.0"
      on Release: ActivateScreen("System settings", 0)
   Button "HmiScreenItemData_2" at 36,213 size 159x47; TextOff 'System information'; PictureOff "Navigates to System information for TP1200 Comfort 16.0.0.0"; PictureOn "Navigates to System information for TP1200 Comfort 16.0.0.0"
      on Release: ActivateScreen("System information", 0)

screen "SIMATIC PLC system diagnostics" 1280x740, template "Template_1"
   on GenerateScreen: SetTag("Tag_ScreenNumber", 6)
   SysDiagControl "HmiScreenItemData" at 1,49 size 1276x623
   Button "Back" at 1,1 size 159x47; TextOff 'Back'
      on Release: ActivateScreen("System screens", 0)

screen "System settings" 1280x740, template "Template_1"
   on GenerateScreen: SetTag("Tag_ScreenNumber", 7)
   Button "Calibrate screen" at 36,95 size 159x47; TextOff 'Calibrate screen'
      on Release: function_bc3e350c()
   Button "Clean screen" at 36,154 size 159x47; TextOff 'Clean screen'
      on Release: function_be740847(30)
   Button "Back" at 1,1 size 159x47; TextOff 'Back'
      on Release: ActivateScreen("System screens", 0)

screen "System information" 1280x740, template "Template_1"
   on GenerateScreen: SetTag("Tag_ScreenNumber", 8)
   TextField "HmiScreenItemData" at 35,51 size 171x28; Text 'HMI device type:'
   TextField "HmiScreenItemData_1" at 241,51 size 1004x28; Text 'TP1200 Comfort 16.0.0.0'
   TextField "HmiScreenItemData_2" at 35,81 size 171x28; Text 'Version:'
   TextField "HmiScreenItemData_3" at 35,111 size 171x28; Text 'Connection:'
   TextField "HmiScreenItemData_4" at 241,111 size 1004x28; Text 'ETHERNET'
   TextField "HmiScreenItemData_5" at 35,141 size 171x28; Text 'PLC:'
   TextField "HmiScreenItemData_6" at 241,141 size 1004x28; Text 'SIMATIC S7 1200'
   Button "Display version" at 241,81 size 1004x28; TextOff 'Display version'
      on Release: function_febcb963(-1)
   Button "Back" at 1,1 size 159x47; TextOff 'Back'
      on Release: ActivateScreen("System screens", 0)
*)